REGION Network 32: Positioning commands
   RUNG wire#powerrail
      Contact( #STC_tUSER_DATA.tR.xReadyToMove )
      wire#w1
      Contact( #IN_xRun )
      wire#w2
      Contact( #STC_tOS.x0 )
      wire#w3
      I_Contact( #STC_tPZD_Pos.tW.tPOS_STW1.x12 )
      Coil( #STC_tPZD_Pos.tW.tSTW1.x6 )
   END_RUNG
   RUNG wire#w1
      Contact( #IN_xReverse )
   END_RUNG wire#w2
   RUNG wire#w1
      Contact( #STC_tST.x0 )
      Contact( #IN_xPositioning )
   END_RUNG wire#w2
   RUNG wire#w2
      Contact( #STC_tOS.x1 )
   END_RUNG wire#w3
   RUNG wire#w2
      Contact( #STC_tOS.x6 )
   END_RUNG wire#w3
   RUNG wire#w2
      Contact( #STC_tPH.x1 )
   END_RUNG wire#w3
   RUNG wire#w2
      Contact( #STC_tPH.x3 )
   END_RUNG wire#w3
   RUNG wire#w2
      Contact( #STC_tPH.x5 )
   END_RUNG wire#w3
   RUNG wire#w2
      Contact( #STC_tPZD_Pos.tW.tSTW1.x6 )
      I_Contact( #STC_tPZD_Pos.tR.tZSW1.x12 )
   END_RUNG wire#w3
   RUNG wire#w1
      Contact( #IN_xRun )
      wire#w4
      Coil( #STC_tPZD_Pos.tW.tSTW1.x5 )
   END_RUNG
   RUNG wire#w1
      Contact( #IN_xReverse )
   END_RUNG wire#w4
   RUNG wire#w1
      Contact( #STC_tST.x0 )
      Contact( #IN_xPositioning )
   END_RUNG wire#w4
   RUNG wire#w1
      Contact( #IN_xRun )
      wire#w5
      Coil( #STC_tPZD_Pos.tW.tSTW1.x4 )
   END_RUNG
   RUNG wire#w1
      Contact( #IN_xReverse )
   END_RUNG wire#w5
   RUNG wire#w1
      Contact( #IN_xPositioning )
   END_RUNG wire#w5
   RUNG wire#w1
      Contact( #OUT_xFeedback )
      I_Contact( #STC_tUSER_DATA.tW.xSafetyStop )
   END_RUNG wire#w5
   RUNG wire#w1
      Contact( #STC_tPH.x6 )
      Coil( #STC_tPZD_Pos.tW.tSTW1.x11 )
   END_RUNG
   // the same network as SCL:
   #STC_tPZD_Pos.tW.tSTW1.x6 := #STC_tUSER_DATA.tR.xReadyToMove AND (#IN_xRun OR #IN_xReverse OR (#STC_tST.x0 AND #IN_xPositioning)) AND (#STC_tOS.x0 OR #STC_tOS.x1 OR #STC_tOS.x6 OR #STC_tPH.x1 OR #STC_tPH.x3 OR #STC_tPH.x5 OR (#STC_tPZD_Pos.tW.tSTW1.x6 AND NOT #STC_tPZD_Pos.tR.tZSW1.x12)) AND NOT #STC_tPZD_Pos.tW.tPOS_STW1.x12;
   #STC_tPZD_Pos.tW.tSTW1.x5 := #STC_tUSER_DATA.tR.xReadyToMove AND (#IN_xRun OR #IN_xReverse OR (#STC_tST.x0 AND #IN_xPositioning));
   #STC_tPZD_Pos.tW.tSTW1.x4 := #STC_tUSER_DATA.tR.xReadyToMove AND (#IN_xRun OR #IN_xReverse OR #IN_xPositioning OR (#OUT_xFeedback AND NOT #STC_tUSER_DATA.tW.xSafetyStop));
   #STC_tPZD_Pos.tW.tSTW1.x11 := #STC_tUSER_DATA.tR.xReadyToMove AND #STC_tPH.x6;
END_REGION

REGION Network 33: Choose positioning type
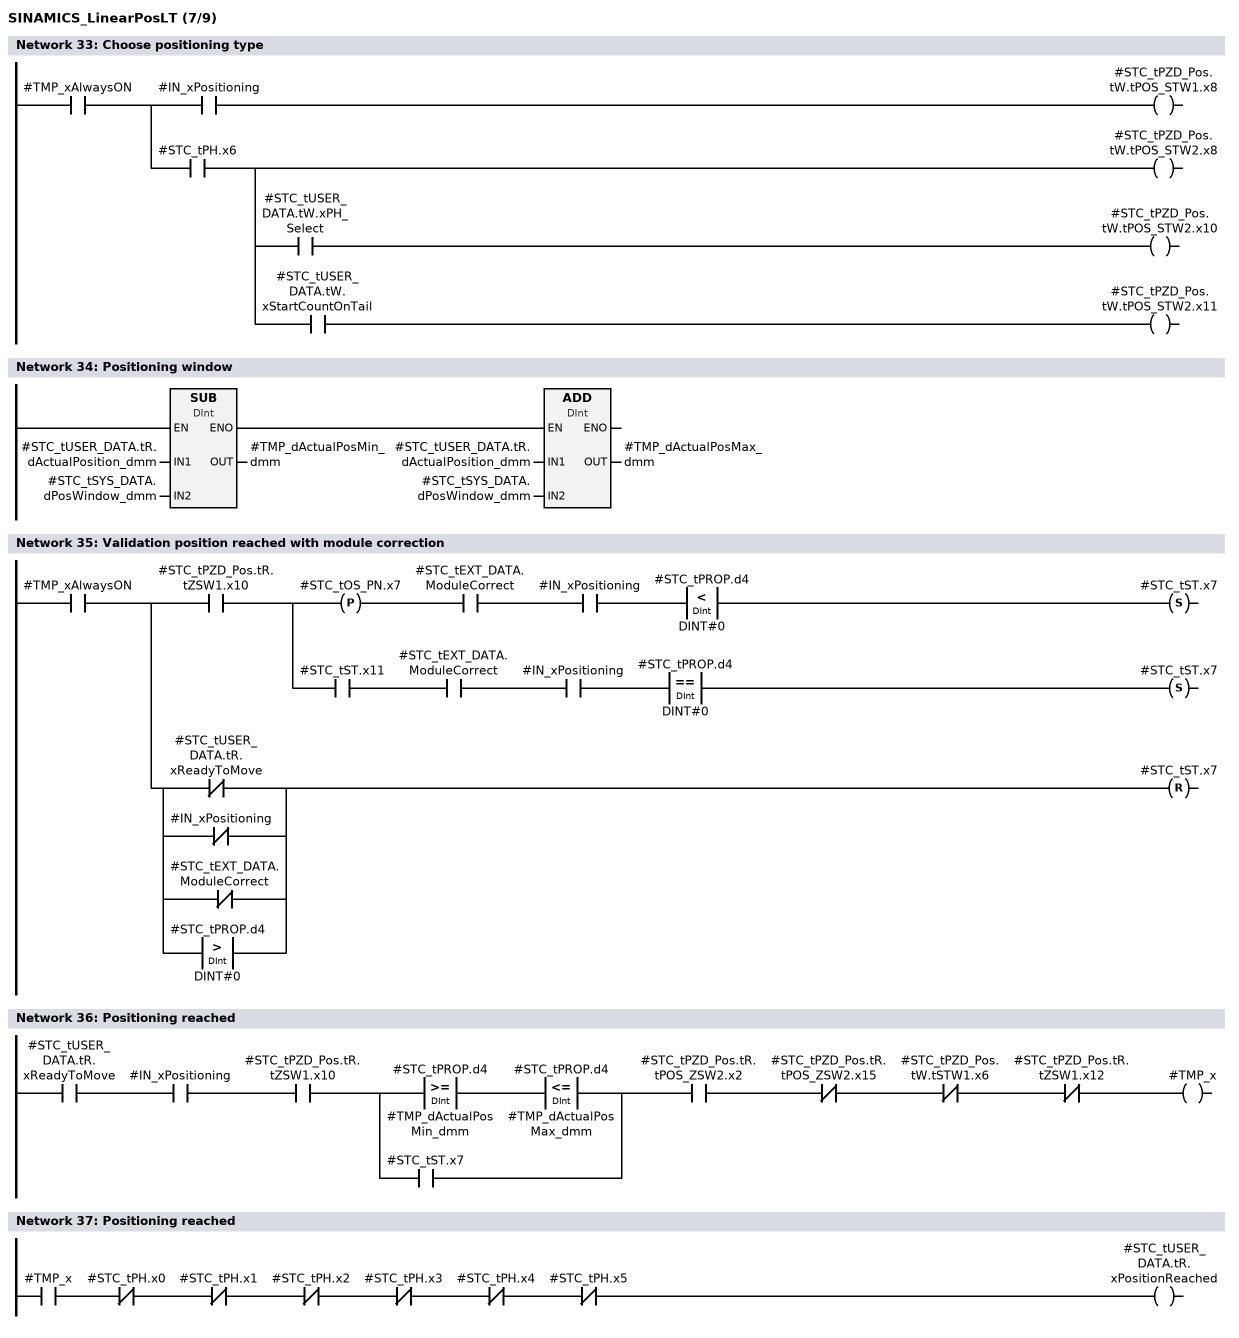
   RUNG wire#powerrail
      Contact( #TMP_xAlwaysON )
      wire#w1
      Contact( #IN_xPositioning )
      Coil( #STC_tPZD_Pos.tW.tPOS_STW1.x8 )
   END_RUNG
   RUNG wire#w1
      Contact( #STC_tPH.x6 )
      wire#w2
      Coil( #STC_tPZD_Pos.tW.tPOS_STW2.x8 )
   END_RUNG
   RUNG wire#w2
      Contact( #STC_tUSER_DATA.tW.xPH_Select )
      Coil( #STC_tPZD_Pos.tW.tPOS_STW2.x10 )
   END_RUNG
   RUNG wire#w2
      Contact( #STC_tUSER_DATA.tW.xStartCountOnTail )
      Coil( #STC_tPZD_Pos.tW.tPOS_STW2.x11 )
   END_RUNG
   // the same network as SCL:
   #STC_tPZD_Pos.tW.tPOS_STW1.x8 := #TMP_xAlwaysON AND #IN_xPositioning;
   #STC_tPZD_Pos.tW.tPOS_STW2.x8 := #TMP_xAlwaysON AND #STC_tPH.x6;
   #STC_tPZD_Pos.tW.tPOS_STW2.x10 := #STC_tPZD_Pos.tW.tPOS_STW2.x8 AND #STC_tUSER_DATA.tW.xPH_Select;
   #STC_tPZD_Pos.tW.tPOS_STW2.x11 := #STC_tPZD_Pos.tW.tPOS_STW2.x8 AND #STC_tUSER_DATA.tW.xStartCountOnTail;
END_REGION

REGION Network 34: Positioning window
   RUNG wire#powerrail
      { S7_Templates := "SrcType := DInt"; S7_GenerateENO := "TRUE" } Sub(in1 := #STC_tUSER_DATA.tR.dActualPosition_dmm, in2 := #STC_tSYS_DATA.dPosWindow_dmm, out => #TMP_dActualPosMin_dmm)
      { S7_Templates := "SrcType := DInt"; S7_GenerateENO := "TRUE" } Add(in1 := #STC_tUSER_DATA.tR.dActualPosition_dmm, in2 := #STC_tSYS_DATA.dPosWindow_dmm, out => #TMP_dActualPosMax_dmm)
   END_RUNG
   // the same network as SCL:
   // ENO of a box is taken as its EN; it also drops when the box reports an error
   #TMP_dActualPosMin_dmm := #STC_tUSER_DATA.tR.dActualPosition_dmm - #STC_tSYS_DATA.dPosWindow_dmm;
   #TMP_dActualPosMax_dmm := #STC_tUSER_DATA.tR.dActualPosition_dmm + #STC_tSYS_DATA.dPosWindow_dmm;
END_REGION

REGION Network 35: Validation position reached with module correction
   RUNG wire#powerrail
      Contact( #TMP_xAlwaysON )
      wire#w1
      Contact( #STC_tPZD_Pos.tR.tZSW1.x10 )
      wire#w2
      P_Trig( #STC_tOS_PN.x7 )
      Contact( #STC_tEXT_DATA.ModuleCorrect )
      Contact( #IN_xPositioning )
      { S7_Templates := "SrcType := DInt" } LT_Contact(in1 := #STC_tPROP.d4, in2 := DINT#0)
      S_Coil( #STC_tST.x7 )
   END_RUNG
   RUNG wire#w2
      Contact( #STC_tST.x11 )
      Contact( #STC_tEXT_DATA.ModuleCorrect )
      Contact( #IN_xPositioning )
      { S7_Templates := "SrcType := DInt" } EQ_Contact(in1 := #STC_tPROP.d4, in2 := DINT#0)
      S_Coil( #STC_tST.x7 )
   END_RUNG
   RUNG wire#w1
      I_Contact( #STC_tUSER_DATA.tR.xReadyToMove )
      wire#w3
      R_Coil( #STC_tST.x7 )
   END_RUNG
   RUNG wire#w1
      I_Contact( #IN_xPositioning )
   END_RUNG wire#w3
   RUNG wire#w1
      I_Contact( #STC_tEXT_DATA.ModuleCorrect )
   END_RUNG wire#w3
   RUNG wire#w1
      { S7_Templates := "SrcType := DInt" } GT_Contact(in1 := #STC_tPROP.d4, in2 := DINT#0)
   END_RUNG wire#w3
   // the same network as SCL:
   #_w1 := #TMP_xAlwaysON AND #STC_tPZD_Pos.tR.tZSW1.x10;
   #_w2 := #_w1 AND NOT #STC_tOS_PN.x7;   // rising edge
   #STC_tOS_PN.x7 := #_w1;
   IF #_w2 AND #STC_tEXT_DATA.ModuleCorrect AND #IN_xPositioning AND (#STC_tPROP.d4 < DINT#0) THEN
       #STC_tST.x7 := TRUE;
   END_IF;
   IF #_w1 AND #STC_tST.x11 AND #STC_tEXT_DATA.ModuleCorrect AND #IN_xPositioning AND (#STC_tPROP.d4 = DINT#0) THEN
       #STC_tST.x7 := TRUE;
   END_IF;
   IF #TMP_xAlwaysON AND (NOT #STC_tUSER_DATA.tR.xReadyToMove OR NOT #IN_xPositioning OR NOT #STC_tEXT_DATA.ModuleCorrect OR (#STC_tPROP.d4 > DINT#0)) THEN
       #STC_tST.x7 := FALSE;
   END_IF;
END_REGION

REGION Network 36: Positioning reached
   RUNG wire#powerrail
      Contact( #STC_tUSER_DATA.tR.xReadyToMove )
      Contact( #IN_xPositioning )
      Contact( #STC_tPZD_Pos.tR.tZSW1.x10 )
      wire#w1
      { S7_Templates := "SrcType := DInt" } GE_Contact(in1 := #STC_tPROP.d4, in2 := #TMP_dActualPosMin_dmm)
      { S7_Templates := "SrcType := DInt" } LE_Contact(in1 := #STC_tPROP.d4, in2 := #TMP_dActualPosMax_dmm)
      wire#w2
      Contact( #STC_tPZD_Pos.tR.tPOS_ZSW2.x2 )
      I_Contact( #STC_tPZD_Pos.tR.tPOS_ZSW2.x15 )
      I_Contact( #STC_tPZD_Pos.tW.tSTW1.x6 )
      I_Contact( #STC_tPZD_Pos.tR.tZSW1.x12 )
      Coil( #TMP_x )
   END_RUNG
   RUNG wire#w1
      Contact( #STC_tST.x7 )
   END_RUNG wire#w2
   // the same network as SCL:
   #TMP_x := #STC_tUSER_DATA.tR.xReadyToMove AND #IN_xPositioning AND #STC_tPZD_Pos.tR.tZSW1.x10 AND (((#STC_tPROP.d4 >= #TMP_dActualPosMin_dmm) AND (#STC_tPROP.d4 <= #TMP_dActualPosMax_dmm)) OR #STC_tST.x7) AND #STC_tPZD_Pos.tR.tPOS_ZSW2.x2 AND NOT #STC_tPZD_Pos.tR.tPOS_ZSW2.x15 AND NOT #STC_tPZD_Pos.tW.tSTW1.x6 AND NOT #STC_tPZD_Pos.tR.tZSW1.x12;
END_REGION

REGION Network 37: Positioning reached
   RUNG wire#powerrail
      Contact( #TMP_x )
      I_Contact( #STC_tPH.x0 )
      I_Contact( #STC_tPH.x1 )
      I_Contact( #STC_tPH.x2 )
      I_Contact( #STC_tPH.x3 )
      I_Contact( #STC_tPH.x4 )
      I_Contact( #STC_tPH.x5 )
      Coil( #STC_tUSER_DATA.tR.xPositionReached )
   END_RUNG
   // the same network as SCL:
   #STC_tUSER_DATA.tR.xPositionReached := #TMP_x AND NOT #STC_tPH.x0 AND NOT #STC_tPH.x1 AND NOT #STC_tPH.x2 AND NOT #STC_tPH.x3 AND NOT #STC_tPH.x4 AND NOT #STC_tPH.x5;
END_REGION

REGION Network 38: Reset count
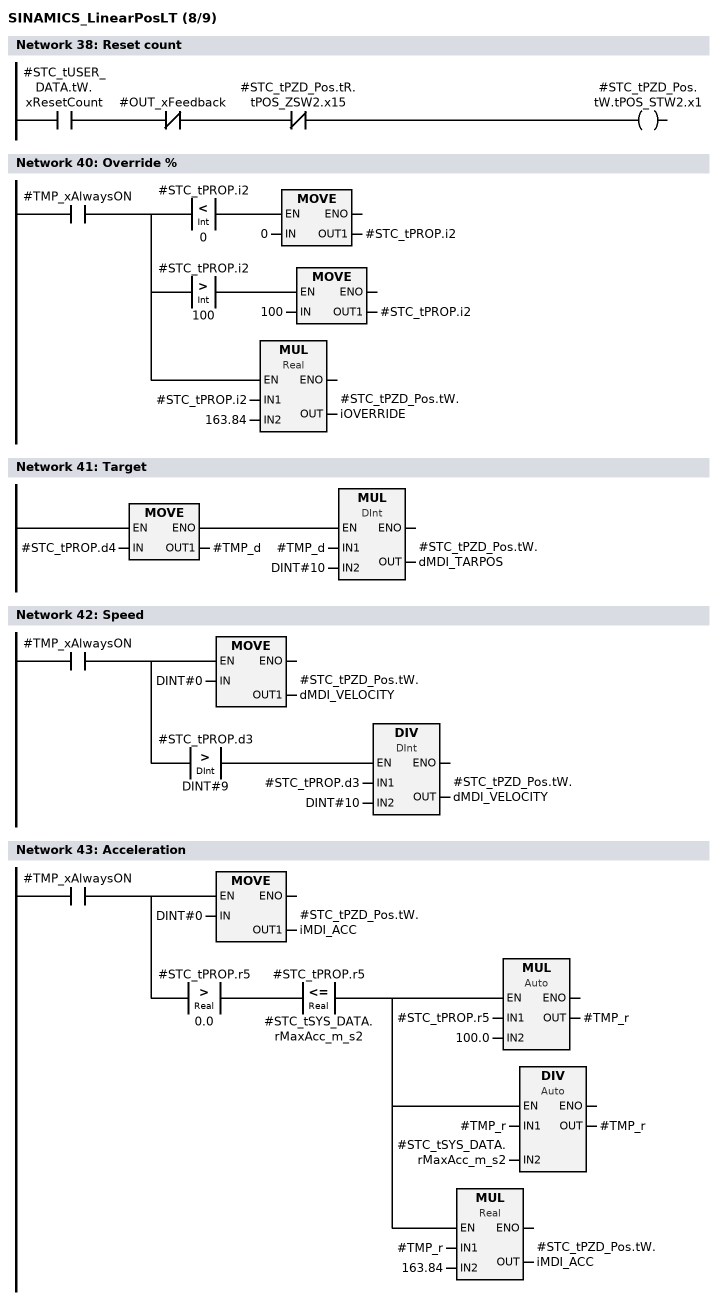
   RUNG wire#powerrail
      Contact( #STC_tUSER_DATA.tW.xResetCount )
      I_Contact( #OUT_xFeedback )
      I_Contact( #STC_tPZD_Pos.tR.tPOS_ZSW2.x15 )
      Coil( #STC_tPZD_Pos.tW.tPOS_STW2.x1 )
   END_RUNG
   // the same network as SCL:
   #STC_tPZD_Pos.tW.tPOS_STW2.x1 := #STC_tUSER_DATA.tW.xResetCount AND NOT #OUT_xFeedback AND NOT #STC_tPZD_Pos.tR.tPOS_ZSW2.x15;
END_REGION

REGION Network 39: #####_PARAMETERS_#####
END_REGION

REGION Network 40: Override %
   RUNG wire#powerrail
      Contact( #TMP_xAlwaysON )
      wire#w1
      { S7_Templates := "SrcType := Int" } LT_Contact(in1 := #STC_tPROP.i2, in2 := 0)
      Move(in := 0, out1 => #STC_tPROP.i2)
   END_RUNG
   RUNG wire#w1
      { S7_Templates := "SrcType := Int" } GT_Contact(in1 := #STC_tPROP.i2, in2 := 100)
      Move(in := 100, out1 => #STC_tPROP.i2)
   END_RUNG
   RUNG wire#w1
      { S7_Templates := "SrcType := Real" } Mul(in1 := #STC_tPROP.i2, in2 := 163.84, out => #STC_tPZD_Pos.tW.iOVERRIDE)
   END_RUNG
   // the same network as SCL:
   IF #TMP_xAlwaysON AND (#STC_tPROP.i2 < 0) THEN #STC_tPROP.i2 := 0; END_IF;
   IF #TMP_xAlwaysON AND (#STC_tPROP.i2 > 100) THEN #STC_tPROP.i2 := 100; END_IF;
   IF #TMP_xAlwaysON THEN #STC_tPZD_Pos.tW.iOVERRIDE := #STC_tPROP.i2 * 163.84; END_IF;
END_REGION

REGION Network 41: Target
   RUNG wire#powerrail
      { S7_GenerateENO := "TRUE" } Move(in := #STC_tPROP.d4, out1 => #TMP_d)
      { S7_Templates := "SrcType := DInt"; S7_GenerateENO := "TRUE" } Mul(in1 := #TMP_d, in2 := DINT#10, out => #STC_tPZD_Pos.tW.dMDI_TARPOS)
   END_RUNG
   // the same network as SCL:
   // ENO of a box is taken as its EN; it also drops when the box reports an error
   #TMP_d := #STC_tPROP.d4;
   #STC_tPZD_Pos.tW.dMDI_TARPOS := #TMP_d * DINT#10;
END_REGION

REGION Network 42: Speed
   RUNG wire#powerrail
      Contact( #TMP_xAlwaysON )
      wire#w1
      { S7_GenerateENO := "TRUE" } Move(in := DINT#0, out1 => #STC_tPZD_Pos.tW.dMDI_VELOCITY)
   END_RUNG
   RUNG wire#w1
      { S7_Templates := "SrcType := DInt" } GT_Contact(in1 := #STC_tPROP.d3, in2 := DINT#9)
      { S7_Templates := "SrcType := DInt"; S7_GenerateENO := "TRUE" } Div(in1 := #STC_tPROP.d3, in2 := DINT#10, out => #STC_tPZD_Pos.tW.dMDI_VELOCITY)
   END_RUNG
   // the same network as SCL:
   IF #TMP_xAlwaysON THEN #STC_tPZD_Pos.tW.dMDI_VELOCITY := DINT#0; END_IF;
   IF #TMP_xAlwaysON AND (#STC_tPROP.d3 > DINT#9) THEN
       #STC_tPZD_Pos.tW.dMDI_VELOCITY := #STC_tPROP.d3 / DINT#10;
   END_IF;
END_REGION

REGION Network 43: Acceleration
   RUNG wire#powerrail
      Contact( #TMP_xAlwaysON )
      wire#w1
      Move(in := DINT#0, out1 => #STC_tPZD_Pos.tW.iMDI_ACC)
   END_RUNG
   RUNG wire#w1
      { S7_Templates := "SrcType := Real" } GT_Contact(in1 := #STC_tPROP.r5, in2 := 0.0)
      { S7_Templates := "SrcType := Real" } LE_Contact(in1 := #STC_tPROP.r5, in2 := #STC_tSYS_DATA.rMaxAcc_m_s2)
      wire#w2
      Mul(in1 := #STC_tPROP.r5, in2 := 100.0, out => #TMP_r)
   END_RUNG
   RUNG wire#w2
      Div(in1 := #TMP_r, in2 := #STC_tSYS_DATA.rMaxAcc_m_s2, out => #TMP_r)
   END_RUNG
   RUNG wire#w2
      { S7_Templates := "SrcType := Real" } Mul(in1 := #TMP_r, in2 := 163.84, out => #STC_tPZD_Pos.tW.iMDI_ACC)
   END_RUNG
   // the same network as SCL:
   IF #TMP_xAlwaysON THEN #STC_tPZD_Pos.tW.iMDI_ACC := DINT#0; END_IF;
   IF #TMP_xAlwaysON AND (#STC_tPROP.r5 > 0.0) AND (#STC_tPROP.r5 <= #STC_tSYS_DATA.rMaxAcc_m_s2) THEN
       #TMP_r := #STC_tPROP.r5 * 100.0;
       #TMP_r := #TMP_r / #STC_tSYS_DATA.rMaxAcc_m_s2;
       #STC_tPZD_Pos.tW.iMDI_ACC := #TMP_r * 163.84;
   END_IF;
END_REGION

REGION Network 44: Deceleration
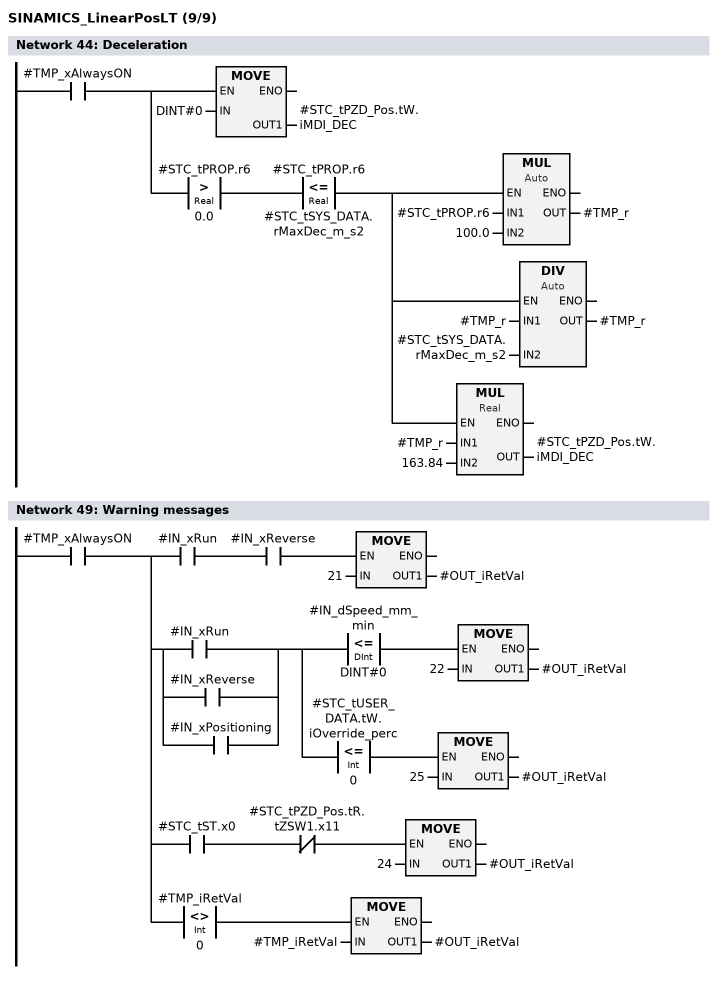
   RUNG wire#powerrail
      Contact( #TMP_xAlwaysON )
      wire#w1
      Move(in := DINT#0, out1 => #STC_tPZD_Pos.tW.iMDI_DEC)
   END_RUNG
   RUNG wire#w1
      { S7_Templates := "SrcType := Real" } GT_Contact(in1 := #STC_tPROP.r6, in2 := 0.0)
      { S7_Templates := "SrcType := Real" } LE_Contact(in1 := #STC_tPROP.r6, in2 := #STC_tSYS_DATA.rMaxDec_m_s2)
      wire#w2
      Mul(in1 := #STC_tPROP.r6, in2 := 100.0, out => #TMP_r)
   END_RUNG
   RUNG wire#w2
      Div(in1 := #TMP_r, in2 := #STC_tSYS_DATA.rMaxDec_m_s2, out => #TMP_r)
   END_RUNG
   RUNG wire#w2
      { S7_Templates := "SrcType := Real" } Mul(in1 := #TMP_r, in2 := 163.84, out => #STC_tPZD_Pos.tW.iMDI_DEC)
   END_RUNG
   // the same network as SCL:
   IF #TMP_xAlwaysON THEN #STC_tPZD_Pos.tW.iMDI_DEC := DINT#0; END_IF;
   IF #TMP_xAlwaysON AND (#STC_tPROP.r6 > 0.0) AND (#STC_tPROP.r6 <= #STC_tSYS_DATA.rMaxDec_m_s2) THEN
       #TMP_r := #STC_tPROP.r6 * 100.0;
       #TMP_r := #TMP_r / #STC_tSYS_DATA.rMaxDec_m_s2;
       #STC_tPZD_Pos.tW.iMDI_DEC := #TMP_r * 163.84;
   END_IF;
END_REGION

REGION Network 45: ################_MOTOR_MODULE_TELEGRAMS_ENDING_#################
END_REGION

REGION Network 46 (STL): Output copy motor module
         L     12;
         T     #TMP_iAddressLength;

   //Compute destination position
         L;
         LAR1;
   //byte 1 = 10h (FIXED for S7)
         L     B#16#10;
         T     B[AR1, P#0.0];
   //byte 2 = data type
         L     B#16#4;  //4 = word
         T     B[AR1, P#1.0];
   //byte 3 & 4 = number of element
         L     #TMP_iAddressLength;  //Production data
         T     W[AR1, P#2.0];
   //byte 5 & 6 = number of DB
         L     0;  //DB production data
         T     W[AR1, P#4.0];
   //byte 7 = memory area
         L     B#16#82;  //82h = Q (Output)
         T     B[AR1, P#6.0];
   //byte 8 & 9 = address. Bit 0,1,2 of tenth byte is bit offset
   //byte 7 = address (high). Valid value = 0-7. Bit 3,4,5,6,7 always 0
         L     #STC_tSYS_DATA.iIOAddress_MM;  //Item size
         SLW   3;
         T     W[AR1, P#8.0];
         SRD   16;
         AW    16#0007;
         T     B[AR1, P#7.0];

         CALL  BLKMOV
         ( SRCBLK  := #STC_tPZD_Pos.tW,
           RET_VAL := #TMP_iRetVal,
           DSTBLK  := #TMP_a
         );
END_REGION

REGION Network 47: #####_RETVAL_RESPONSE_#####
END_REGION

REGION Network 48 (STL): Initialize RetVal
         L     0;
         T     #OUT_iRetVal;
END_REGION

REGION Network 49: Warning messages
   RUNG wire#powerrail
      Contact( #TMP_xAlwaysON )
      wire#w1
      Contact( #IN_xRun )
      Contact( #IN_xReverse )
      Move(in := 21, out1 => #OUT_iRetVal)
   END_RUNG
   RUNG wire#w1
      Contact( #IN_xRun )
      wire#w2
      { S7_Templates := "SrcType := DInt" } LE_Contact(in1 := #IN_dSpeed_mm_min, in2 := DINT#0)
      Move(in := 22, out1 => #OUT_iRetVal)
   END_RUNG
   RUNG wire#w1
      Contact( #IN_xReverse )
   END_RUNG wire#w2
   RUNG wire#w1
      Contact( #IN_xPositioning )
   END_RUNG wire#w2
   RUNG wire#w2
      { S7_Templates := "SrcType := Int" } LE_Contact(in1 := #STC_tUSER_DATA.tW.iOverride_perc, in2 := 0)
      Move(in := 25, out1 => #OUT_iRetVal)
   END_RUNG
   RUNG wire#w1
      Contact( #STC_tST.x0 )
      I_Contact( #STC_tPZD_Pos.tR.tZSW1.x11 )
      Move(in := 24, out1 => #OUT_iRetVal)
   END_RUNG
   RUNG wire#w1
      { S7_Templates := "SrcType := Int" } NE_Contact(in1 := #TMP_iRetVal, in2 := 0)
      Move(in := #TMP_iRetVal, out1 => #OUT_iRetVal)
   END_RUNG
   // the same network as SCL:
   IF #TMP_xAlwaysON AND #IN_xRun AND #IN_xReverse THEN #OUT_iRetVal := 21; END_IF;
   #_w1 := #TMP_xAlwaysON AND (#IN_xRun OR #IN_xReverse OR #IN_xPositioning);
   IF #_w1 AND (#IN_dSpeed_mm_min <= DINT#0) THEN #OUT_iRetVal := 22; END_IF;
   IF #_w1 AND (#STC_tUSER_DATA.tW.iOverride_perc <= 0) THEN #OUT_iRetVal := 25; END_IF;
   IF #TMP_xAlwaysON AND #STC_tST.x0 AND NOT #STC_tPZD_Pos.tR.tZSW1.x11 THEN #OUT_iRetVal := 24; END_IF;
   IF #TMP_xAlwaysON AND (#TMP_iRetVal <> 0) THEN #OUT_iRetVal := #TMP_iRetVal; END_IF;
END_REGION

REGION Network 50 (STL): Blocking messages
         JU    Rest;
   Err:  T     #OUT_iRetVal;
END_REGION

REGION Network 51 (STL): Reset input commands
   // R     #USER_DATA.W.SafetyStop
   //       R     #USER_DATA.W.FlyChange
   //       R     #USER_DATA.W.PH_Select
   //       R     #USER_DATA.W.StartCountOnHead
   //       R     #USER_DATA.W.StartCountOnTail
   //       R     #USER_DATA.W.BrakeRelease
   //       R     #USER_DATA.W.ResetCount
   //       R     #USER_DATA.W.PresetRq
   //       R     #USER_DATA.W.HomeSearch
   //       R     #USER_DATA.W.ReverseHoming
   //       R     #USER_DATA.W.ReferenceCam
   //       R     #USER_DATA.W.ReferenceZero
   //       R     #USER_DATA.W.MDI_Continue
   //       R     #USER_DATA.W.SwLimitsEnable
   //       R     #USER_DATA.W.HwLimitsEnable
   //       R     #Run
   //       R     #Reverse
   //       R     #Positioning
   // 
   //       L     L#0
   //       T     #Speed
   //       T     #USER_DATA.W.Override
   //       T     #USER_DATA.W.Target
   //       T     #USER_DATA.W.Preset
   //       T     #USER_DATA.W.Acc
   //       T     #USER_DATA.W.Dec
   Rest: NOP   0;
   //    SET
   //    R     #IN_xDrive_EN
   //    R     #IN_xResetFaults
END_REGION

REGION Network 52 (STL): Restore AR1 & AR2 value
   //    L     #TMP_dOldValue_AR1
   //    LAR1
   //    L     #TMP_dOldValue_AR2
   //    LAR2
END_REGION
END_FUNCTION_BLOCK

FUNCTION_BLOCK "SINAMICS_Rotator"   // FB55, LAD
TITLE = Sinamics drive manager
{ S7_Optimized_Access := 'FALSE' }
AUTHOR : Armitano
VERSION : 1.4
// Return value:
// * 0: OK
// Blocking message:
// * group 1 to 9: general error
// * group 10 to 19: system data error
//   * 10: Sinamics input/output addresses wrong or not setted
//   * 11: Maximum speed in Rpm wrong or not setted
//   * 13: Conversion coefficent for rpm to °/min wrong or not setted
//   * 14: Maximum acceleration wrong or not setted
//   * 15: Maximum deceleration wrong or not setted
// Warning message:
// * group 20 to 29: user data error
//   * 21: Run command + reverse command no possixle
//   * 22: Preset speed at zero during run/reverse command
//   * 24: Axes no referenced
// Other:
// * group 30 to 32: preset data error
//   * 30: Error during send preset value (Check parameters in Sys_Data)
//   * 31: Error during preset command (Check parameters in Sys_Data)
//   * 32: Error during saving preset command (Check Sys_Data)
//   * 34: Error during send preset homing (Check parameters in Sys_Data)
// * group 8000 to 9000: SFC20 code (Read the SFC20 Help)
   VAR_INPUT
      IN_xDrive_EN : Bool;   // Drive enable
      IN_xRun : Bool;   // Run clockwise
      IN_xReverse : Bool;   // Run counterclockwise
      IN_xResetFaults : Bool;   // Reset faults
      IN_dSpeed_deg_min : DInt;   // Speed reference [°/min]
   END_VAR
   VAR_OUTPUT
      OUT_xFeedback : Bool;   // Feedback active
      OUT_xFaultPresent : Bool;   // Fault present
      OUT_iFaultCode : Int;   // Fault code
      OUT_iRetVal : Int;   // Return value in case of wrong configuration
   END_VAR
   VAR
      STC_tUSER_DATA : Struct   // User data (Extended functions commands for execute the application desired)
         tR : Struct
            xReadyfForSwitchOn : Bool;   // Ready for switch on
            xReadyToMove : Bool;   // Ready to move
            xAxleRefered : Bool;   // Axle referenced
            xPositionReached : Bool;   // Position reached
            xAlarmPresent : Bool;   // Alarm present
            iAlarmCode : Int;   // Alarm code
            dActualPosition_cdeg : DInt;   // Actual position value [°/100]
            dActualSpeed_deg_min : DInt;   // Actual speed value [°/min]
         END_STRUCT;
         tW : Struct
            xSafetyStop : Bool;   // Safety stop (OFF3)
            x2 : Bool;
            xJogMode : Bool;   // Jog modality (Free movment)
            x4 : Bool;
            x5 : Bool;
            xBrakeRelease : Bool;   // Brake release
            x7 : Bool;
            xPresetRq : Bool;   // Preset request
            x9 : Bool;
            x10 : Bool;
            x11 : Bool;
            x12 : Bool;
            x13 : Bool;
            x14 : Bool;
            x15 : Bool;
            i12 : Int := 100;
            d13 : DInt;
            d14 : DInt;
            rAcc_deg_s2 : Real;   // Acceleration [°/s2]
            rDec_deg_s2 : Real;   // Deceleration [°/s2]
         END_STRUCT;
      END_STRUCT;
      STC_tSYS_DATA : Struct   // System data (Info about applications type and HW config.)
         iIOAddress_MM : Int := -1;   // Input/Output addresses for motor module
         i2 : Int;
         i3 : Int;
         iDiagAddress : Int;   // Diagnostic address of SINAMICS module
         iPosPZD_CU : Int;   // Number of PZD position in SINAMICS configuration [1,2,3..]
         iPosPZD_MM : Int;   // Number of PZD position in SINAMICS configuration [1,2,3..]
         i7 : Int;
         dMaxSpeed_rpm : DInt;   // MaxSpeed [rpm]
         d9 : DInt;
         dPosWindow_cdeg : DInt := L#40;   // Positioning window [°/100]
         d11 : DInt;
         d12 : DInt;
         d13 : DInt;
         rK_rpm_grdMin : Real;   // K Conversion from rpm to °/min
         r15 : Real;
         rMaxAcc_deg_s2 : Real;   // MaxAcc [°/s2]
         rMaxDec_deg_s2 : Real;   // MaxDec [°/s2]
         r18 : Real;
         r19 : Real;
      END_STRUCT;
      STC_tST : Struct
         x0 : Bool;
         x1 : Bool;   // Delay restart positioning
         x2 : Bool;
         x3 : Bool;
         x4 : Bool;
         x5 : Bool;
         x6 : Bool;   // Target = Feedback target
         x7 : Bool;
         x8 : Bool;   // Preset phases in progress
         x9 : Bool;
         x10 : Bool;
         x11 : Bool;
         x12 : Bool;
         x13 : Bool;
         x14 : Bool;
         x15 : Bool;
      END_STRUCT;
      STC_tOS_PN : Struct
         x0 : Bool;   // Run
         x1 : Bool;   // Reverse
         x2 : Bool;
         x3 : Bool;
         x4 : Bool;
         x5 : Bool;
         x6 : Bool;
         x7 : Bool;   // Position reached
         x8 : Bool;
         x9 : Bool;
         x10 : Bool;   // Preset position
         x11 : Bool;
         x12 : Bool;
         x13 : Bool;
         x14 : Bool;
         x15 : Bool;
      END_STRUCT;
      STC_tOS : Struct
         x0 : Bool;   // Run
         x1 : Bool;   // Reverse
         x2 : Bool;
         x3 : Bool;
         x4 : Bool;
         x5 : Bool;
         x6 : Bool;
         x7 : Bool;
         x8 : Bool;
         x9 : Bool;
         x10 : Bool;
         x11 : Bool;
         x12 : Bool;
         x13 : Bool;
         x14 : Bool;
         x15 : Bool;
      END_STRUCT;
      STC_tPH : Struct
         x0 : Bool;   // Positioning initializing
         x1 : Bool;   // Positioning request
         x2 : Bool;
         x3 : Bool;
         x4 : Bool;
         x5 : Bool;
         x6 : Bool;
         x7 : Bool;
         x8 : Bool;   // Send encoder value
         x9 : Bool;
         x10 : Bool;   // Send preset command
         x11 : Bool;
         x12 : Bool;   // Send saving preset command
         x13 : Bool;
         x14 : Bool;   // End preset encoder
         x15 : Bool;
      END_STRUCT;
      STC_tPROP : Struct
         i0 : Int;   // Previous cycle [ms]
         tmON_DelayRestart_ms : IEC_TIMER;   // Delay restart positioning [ms]
         i2 : Int;
         i3 : Int;
         i4 : Int;
         dPulsePos_0_cdeg : DInt;   // Position to 0° [°/100]
         dPulsePos_90_cdeg : DInt := L#9000;   // Position to 90° [°/100]
         dPulsePos_180_cdeg : DInt := L#18000;   // Position to 180° [°/100]
         dPulsePos_270_cdeg : DInt := L#27000;   // Position to 270° [°/100]
      END_STRUCT;
      STC_tMngSysReg : Struct   // Managment system register
         tST : Struct
            xWrite_Request : Bool;
            xDone : Bool;
            xBusy : Bool;
            xError : Bool;
            xSpare4 : Bool;
            xSpare5 : Bool;
            xSpare6 : Bool;
            xSpare7 : Bool;
            ID : Hw_Io;
            dINDEX : DInt;
            uiLEN : UInt;
            dwSTATUS : DWord;
            iSpare : Int;
         END_STRUCT;
         tDATA : Struct
            wRequest_refere_RequestID : Word := W#16#102;   // (Request_referece=01 Alwais=01 )*(RequestID=02 Change Param)
            wAxis_NoOfParameters : Word := W#16#101;   // (Axis=Num.Object)(NoOfParameters=Num of parameter to change)
            wAttribute_NoOfElements : Word := W#16#1001;   // (Attribute=10 Alwais=10)(NoOfParameters=Num of subparameter to Write)
            iParameter_number : Int := 2599;   // Parameter_number=Number of the parameter
            wSubindex : Word;   // Subindex
            wFormat_NoOfValue : Word := W#16#4301;   // (Format_NoOfValue=Format 42=Word 43=Dword)(Num. of value to transfer)
            dwRegisterValue : DWord := DW#16#1;   // Register value
         END_STRUCT;
      END_STRUCT;
      STC_tWriteRecord : WRREC;
      STC_tPZD_Pos : Struct   // Motor module positioner telegram 111
         tR : Struct   // READ
            tZSW1 : Struct   // R2089[0].STATUS WORD 1
               x8 : Bool;   // Tracking error in tolerance
               x9 : Bool;   // Control request
               x10 : Bool;   // Target position reached
               x11 : Bool;   // Reference point set
               x12 : Bool;   // Acknowledgment, travering block activated
               x13 : Bool;   // In_actl < speed threshold value 3
               x14 : Bool;   // Axis accelerating
               x15 : Bool;   // Axis decelerating
               x0 : Bool;   // Ready for switch on
               x1 : Bool;   // Ready
               x2 : Bool;   // Operation enabled
               x3 : Bool;   // Fault present
               x4 : Bool;   // OFF2
               x5 : Bool;   // OFF3
               x6 : Bool;   // Switching on inhibited active
               x7 : Bool;   // Alarm present
            END_STRUCT;
            tPOS_ZSW1 : Struct   // R2089[3].POSITIONER STATUS WORD 2
               x8 : Bool;   // STOP cam minus active
               x9 : Bool;   // STOP cam plus active
               x10 : Bool;   // Jog active
               x11 : Bool;   // Homing procedure active
               x12 : Bool;   // Flying referencing active
               x13 : Bool;   // Traversing block active
               x14 : Bool;   // Setup active
               x15 : Bool;   // MDI active
               x0 : Bool;   // Active traversing block, bit 0
               x1 : Bool;   // Active traversing block, bit 1
               x2 : Bool;   // Active traversing block, bit 2
               x3 : Bool;   // Active traversing block, bit 3
               x4 : Bool;   // Active traversing block, bit 4
               x5 : Bool;   // Active traversing block, bit 5
               x6 : Bool;   // Reserved
               x7 : Bool;   // Reserved
            END_STRUCT;
            tPOS_ZSW2 : Struct   // R2089[4].POSITIONER STATUS WORD 3
               x8 : Bool;   // Position actual value <= cam switching position 1
               x9 : Bool;   // Position actual value <= cam switching position 2